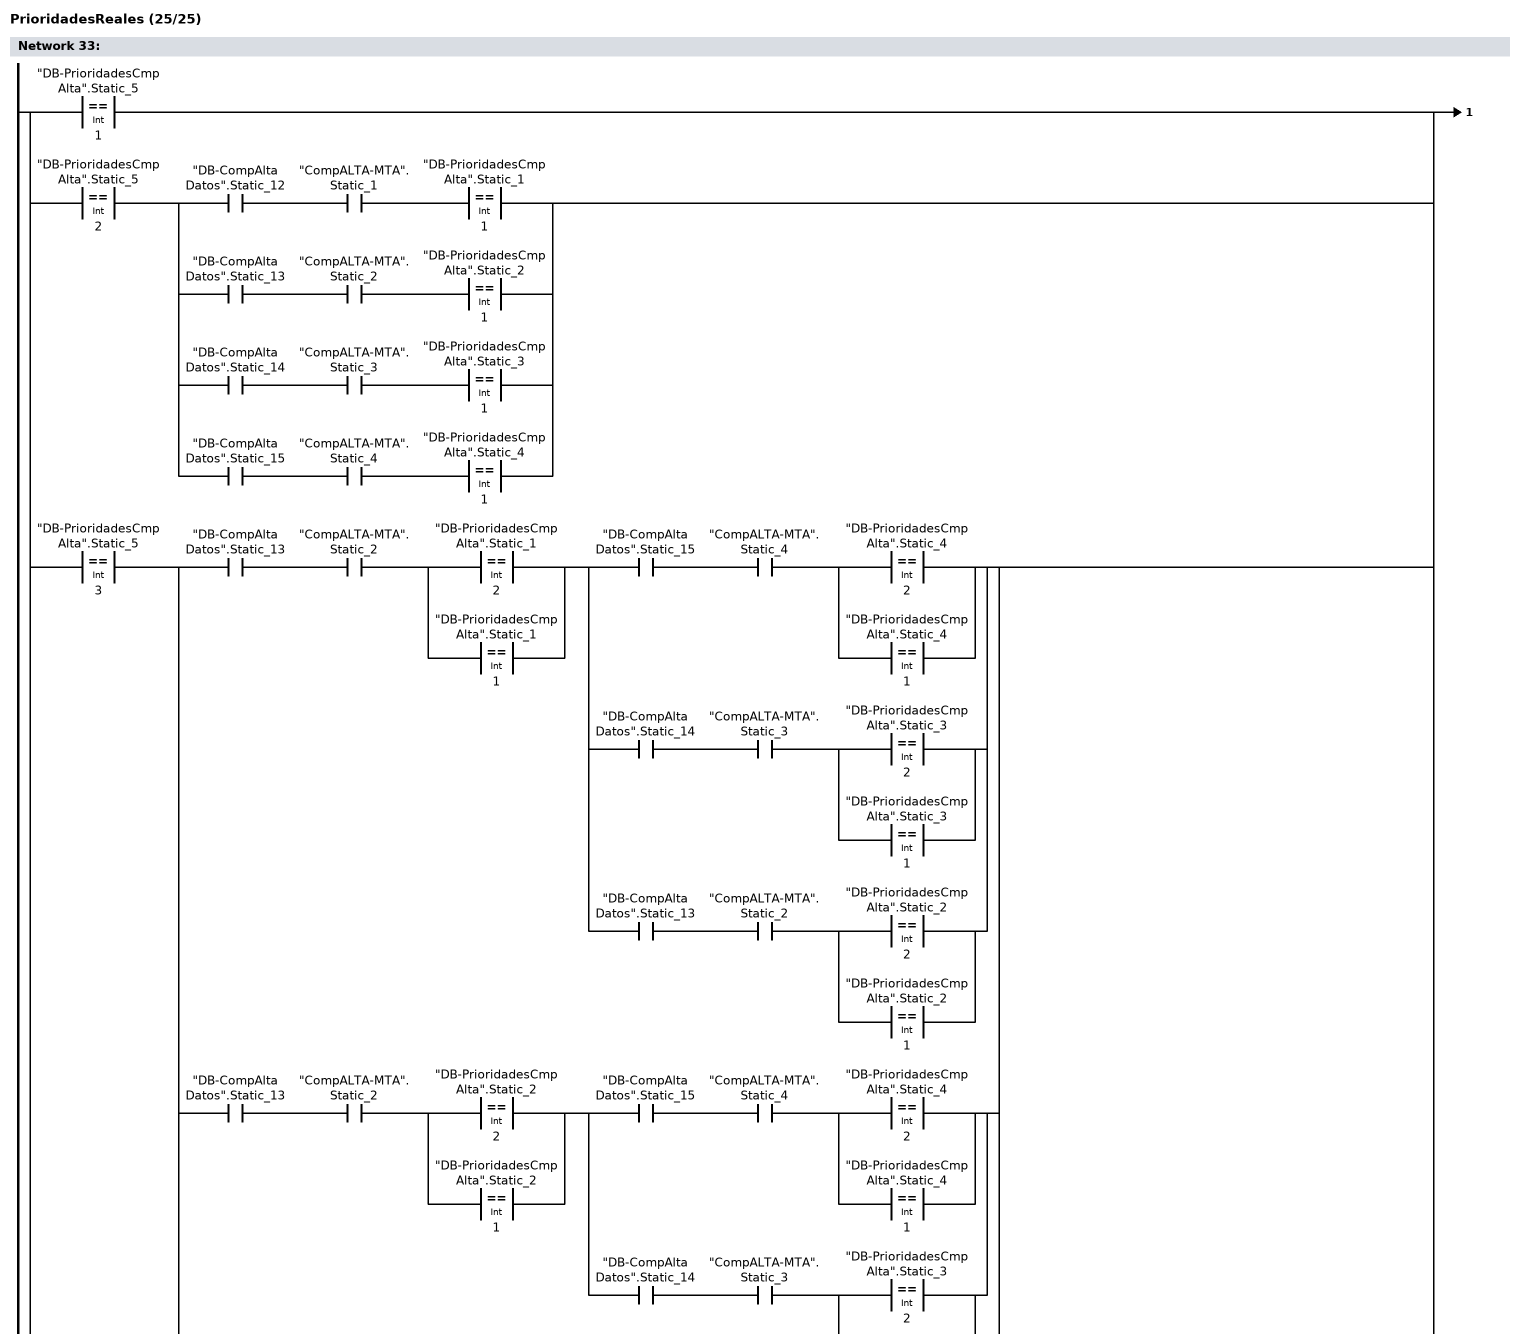
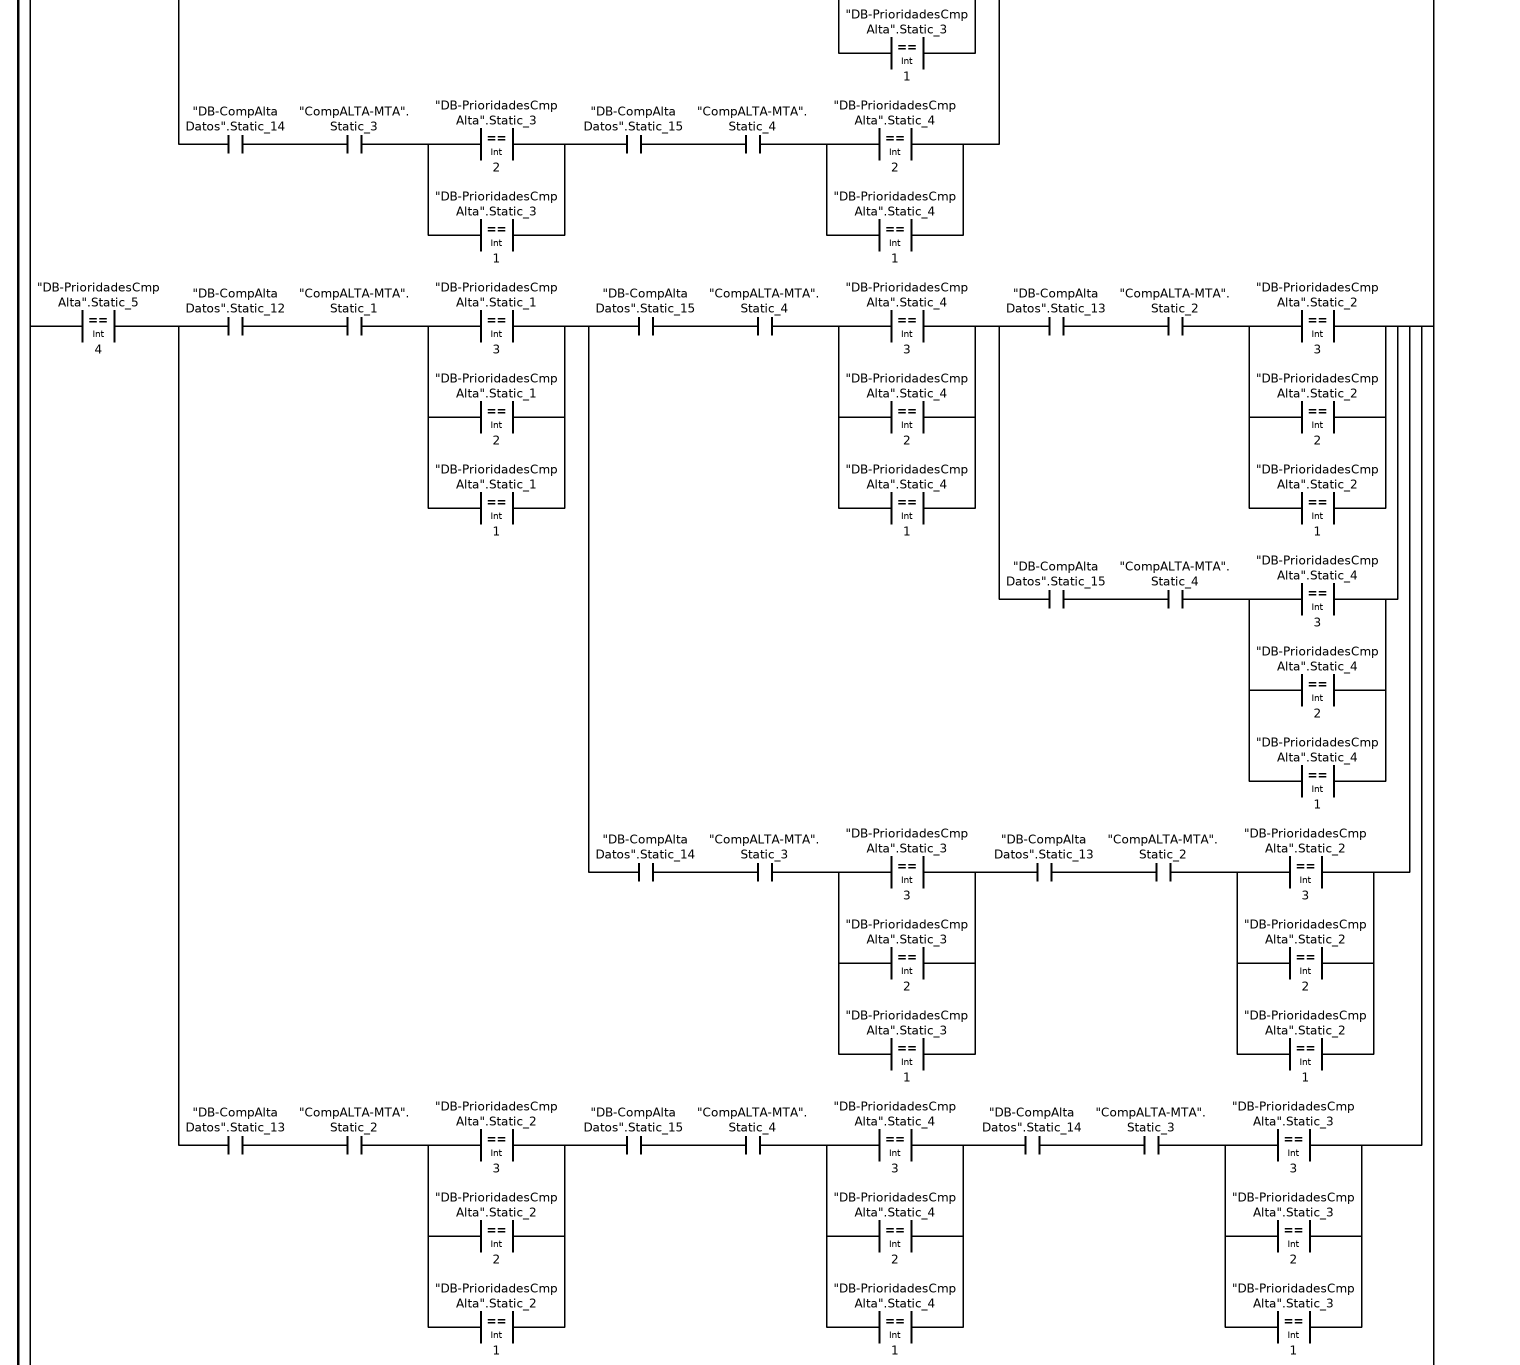
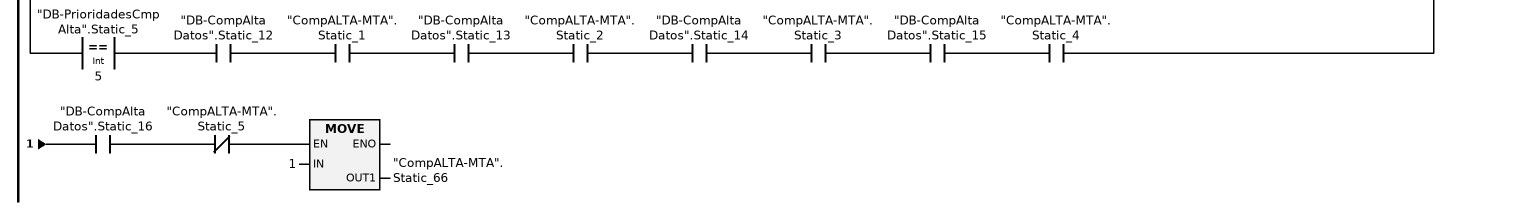
   IF (("DB-PrioridadesCmpAlta".Static_5 = 1) OR (("DB-PrioridadesCmpAlta".Static_5 = 2) AND (("DB-CompAltaDatos".Static_12 AND "CompALTA-MTA".Static_1 AND ("DB-PrioridadesCmpAlta".Static_1 = 1)) OR ("DB-CompAltaDatos".Static_13 AND "CompALTA-MTA".Static_2 AND ("DB-PrioridadesCmpAlta".Static_2 = 1)) OR ("DB-CompAltaDatos".Static_14 AND "CompALTA-MTA".Static_3 AND ("DB-PrioridadesCmpAlta".Static_3 = 1)) OR ("DB-CompAltaDatos".Static_15 AND "CompALTA-MTA".Static_4 AND ("DB-PrioridadesCmpAlta".Static_4 = 1)))) OR (("DB-PrioridadesCmpAlta".Static_5 = 3) AND (("DB-CompAltaDatos".Static_13 AND "CompALTA-MTA".Static_2 AND (("DB-PrioridadesCmpAlta".Static_1 = 2) OR ("DB-PrioridadesCmpAlta".Static_1 = 1)) AND (("DB-CompAltaDatos".Static_15 AND "CompALTA-MTA".Static_4 AND (("DB-PrioridadesCmpAlta".Static_4 = 2) OR ("DB-PrioridadesCmpAlta".Static_4 = 1))) OR ("DB-CompAltaDatos".Static_14 AND "CompALTA-MTA".Static_3 AND (("DB-PrioridadesCmpAlta".Static_3 = 2) OR ("DB-PrioridadesCmpAlta".Static_3 = 1))) OR ("DB-CompAltaDatos".Static_13 AND "CompALTA-MTA".Static_2 AND (("DB-PrioridadesCmpAlta".Static_2 = 2) OR ("DB-PrioridadesCmpAlta".Static_2 = 1))))) OR ("DB-CompAltaDatos".Static_13 AND "CompALTA-MTA".Static_2 AND (("DB-PrioridadesCmpAlta".Static_2 = 2) OR ("DB-PrioridadesCmpAlta".Static_2 = 1)) AND (("DB-CompAltaDatos".Static_15 AND "CompALTA-MTA".Static_4 AND (("DB-PrioridadesCmpAlta".Static_4 = 2) OR ("DB-PrioridadesCmpAlta".Static_4 = 1))) OR ("DB-CompAltaDatos".Static_14 AND "CompALTA-MTA".Static_3 AND (("DB-PrioridadesCmpAlta".Static_3 = 2) OR ("DB-PrioridadesCmpAlta".Static_3 = 1))))) OR ("DB-CompAltaDatos".Static_14 AND "CompALTA-MTA".Static_3 AND (("DB-PrioridadesCmpAlta".Static_3 = 2) OR ("DB-PrioridadesCmpAlta".Static_3 = 1)) AND "DB-CompAltaDatos".Static_15 AND "CompALTA-MTA".Static_4 AND (("DB-PrioridadesCmpAlta".Static_4 = 2) OR ("DB-PrioridadesCmpAlta".Static_4 = 1))))) OR (("DB-PrioridadesCmpAlta".Static_5 = 4) AND (("DB-CompAltaDatos".Static_12 AND "CompALTA-MTA".Static_1 AND (("DB-PrioridadesCmpAlta".Static_1 = 3) OR ("DB-PrioridadesCmpAlta".Static_1 = 2) OR ("DB-PrioridadesCmpAlta".Static_1 = 1)) AND (("DB-CompAltaDatos".Static_15 AND "CompALTA-MTA".Static_4 AND (("DB-PrioridadesCmpAlta".Static_4 = 3) OR ("DB-PrioridadesCmpAlta".Static_4 = 2) OR ("DB-PrioridadesCmpAlta".Static_4 = 1)) AND (("DB-CompAltaDatos".Static_13 AND "CompALTA-MTA".Static_2 AND (("DB-PrioridadesCmpAlta".Static_2 = 3) OR ("DB-PrioridadesCmpAlta".Static_2 = 2) OR ("DB-PrioridadesCmpAlta".Static_2 = 1))) OR ("DB-CompAltaDatos".Static_15 AND "CompALTA-MTA".Static_4 AND (("DB-PrioridadesCmpAlta".Static_4 = 3) OR ("DB-PrioridadesCmpAlta".Static_4 = 2) OR ("DB-PrioridadesCmpAlta".Static_4 = 1))))) OR ("DB-CompAltaDatos".Static_14 AND "CompALTA-MTA".Static_3 AND (("DB-PrioridadesCmpAlta".Static_3 = 3) OR ("DB-PrioridadesCmpAlta".Static_3 = 2) OR ("DB-PrioridadesCmpAlta".Static_3 = 1)) AND "DB-CompAltaDatos".Static_13 AND "CompALTA-MTA".Static_2 AND (("DB-PrioridadesCmpAlta".Static_2 = 3) OR ("DB-PrioridadesCmpAlta".Static_2 = 2) OR ("DB-PrioridadesCmpAlta".Static_2 = 1))))) OR ("DB-CompAltaDatos".Static_13 AND "CompALTA-MTA".Static_2 AND (("DB-PrioridadesCmpAlta".Static_2 = 3) OR ("DB-PrioridadesCmpAlta".Static_2 = 2) OR ("DB-PrioridadesCmpAlta".Static_2 = 1)) AND "DB-CompAltaDatos".Static_15 AND "CompALTA-MTA".Static_4 AND (("DB-PrioridadesCmpAlta".Static_4 = 3) OR ("DB-PrioridadesCmpAlta".Static_4 = 2) OR ("DB-PrioridadesCmpAlta".Static_4 = 1)) AND "DB-CompAltaDatos".Static_14 AND "CompALTA-MTA".Static_3 AND (("DB-PrioridadesCmpAlta".Static_3 = 3) OR ("DB-PrioridadesCmpAlta".Static_3 = 2) OR ("DB-PrioridadesCmpAlta".Static_3 = 1))))) OR (("DB-PrioridadesCmpAlta".Static_5 = 5) AND "DB-CompAltaDatos".Static_12 AND "CompALTA-MTA".Static_1 AND "DB-CompAltaDatos".Static_13 AND "CompALTA-MTA".Static_2 AND "DB-CompAltaDatos".Static_14 AND "CompALTA-MTA".Static_3 AND "DB-CompAltaDatos".Static_15 AND "CompALTA-MTA".Static_4)) AND "DB-CompAltaDatos".Static_16 AND NOT "CompALTA-MTA".Static_5 THEN
       "CompALTA-MTA".Static_66 := 1;
   END_IF;
END_REGION
END_FUNCTION

FUNCTION "FlancosCmpAlta" : Void   // FC45, LAD
{ S7_Optimized_Access := 'FALSE' }
VERSION : 0.1
   VAR_TEMP   // added for the SCL form of the ladder/FBD networks
      _w1 : Bool;
      _w2 : Bool;
      _w3 : Bool;
      _w4 : Bool;
      _w5 : Bool;
      _w6 : Bool;
      _w7 : Bool;
      _s5time1 : S5Time;
   END_VAR
BEGIN

REGION Network 1
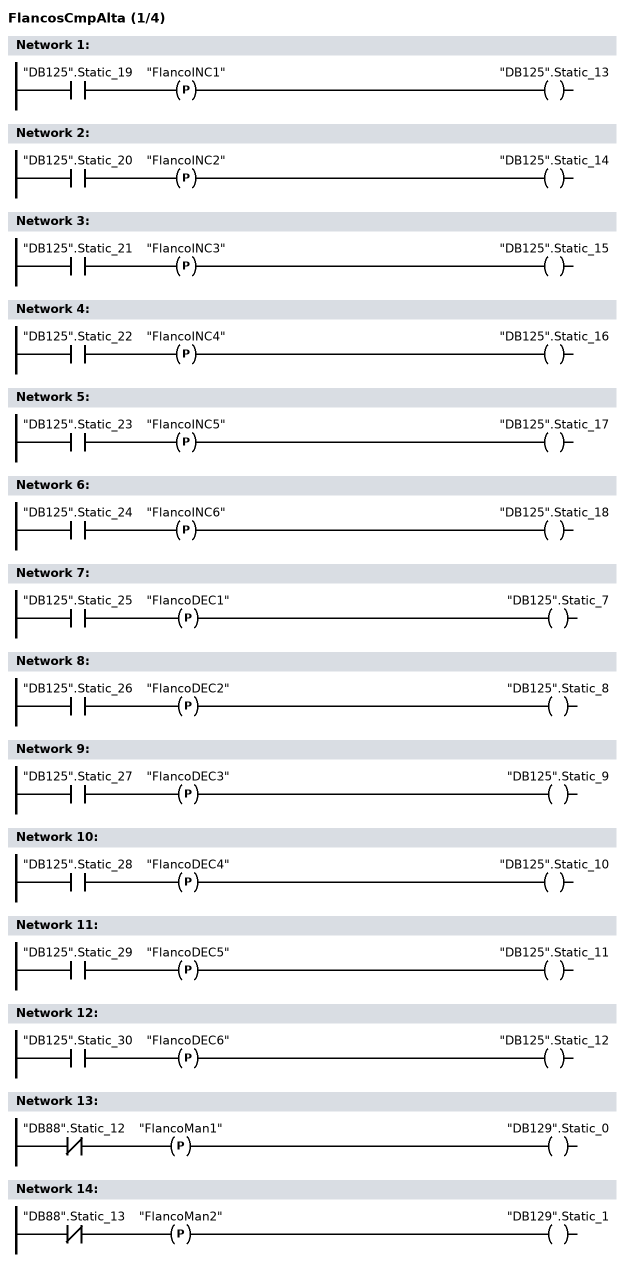
   RUNG wire#powerrail
      Contact( "DB125".Static_19 )
      P_Trig( "FlancoINC1" )
      Coil( "DB125".Static_13 )
   END_RUNG
   // the same network as SCL:
   #_w1 := "DB125".Static_19 AND NOT "FlancoINC1";   // rising edge
   "FlancoINC1" := "DB125".Static_19;
   "DB125".Static_13 := #_w1;
END_REGION

REGION Network 2
   RUNG wire#powerrail
      Contact( "DB125".Static_20 )
      P_Trig( "FlancoINC2" )
      Coil( "DB125".Static_14 )
   END_RUNG
   // the same network as SCL:
   #_w1 := "DB125".Static_20 AND NOT "FlancoINC2";   // rising edge
   "FlancoINC2" := "DB125".Static_20;
   "DB125".Static_14 := #_w1;
END_REGION

REGION Network 3
   RUNG wire#powerrail
      Contact( "DB125".Static_21 )
      P_Trig( "FlancoINC3" )
      Coil( "DB125".Static_15 )
   END_RUNG
   // the same network as SCL:
   #_w1 := "DB125".Static_21 AND NOT "FlancoINC3";   // rising edge
   "FlancoINC3" := "DB125".Static_21;
   "DB125".Static_15 := #_w1;
END_REGION

REGION Network 4
   RUNG wire#powerrail
      Contact( "DB125".Static_22 )
      P_Trig( "FlancoINC4" )
      Coil( "DB125".Static_16 )
   END_RUNG
   // the same network as SCL:
   #_w1 := "DB125".Static_22 AND NOT "FlancoINC4";   // rising edge
   "FlancoINC4" := "DB125".Static_22;
   "DB125".Static_16 := #_w1;
END_REGION

REGION Network 5
   RUNG wire#powerrail
      Contact( "DB125".Static_23 )
      P_Trig( "FlancoINC5" )
      Coil( "DB125".Static_17 )
   END_RUNG
   // the same network as SCL:
   #_w1 := "DB125".Static_23 AND NOT "FlancoINC5";   // rising edge
   "FlancoINC5" := "DB125".Static_23;
   "DB125".Static_17 := #_w1;
END_REGION

REGION Network 6
   RUNG wire#powerrail
      Contact( "DB125".Static_24 )
      P_Trig( "FlancoINC6" )
      Coil( "DB125".Static_18 )
   END_RUNG
   // the same network as SCL:
   #_w1 := "DB125".Static_24 AND NOT "FlancoINC6";   // rising edge
   "FlancoINC6" := "DB125".Static_24;
   "DB125".Static_18 := #_w1;
END_REGION

REGION Network 7
   RUNG wire#powerrail
      Contact( "DB125".Static_25 )
      P_Trig( "FlancoDEC1" )
      Coil( "DB125".Static_7 )
   END_RUNG
   // the same network as SCL:
   #_w1 := "DB125".Static_25 AND NOT "FlancoDEC1";   // rising edge
   "FlancoDEC1" := "DB125".Static_25;
   "DB125".Static_7 := #_w1;
END_REGION

REGION Network 8
   RUNG wire#powerrail
      Contact( "DB125".Static_26 )
      P_Trig( "FlancoDEC2" )
      Coil( "DB125".Static_8 )
   END_RUNG
   // the same network as SCL:
   #_w1 := "DB125".Static_26 AND NOT "FlancoDEC2";   // rising edge
   "FlancoDEC2" := "DB125".Static_26;
   "DB125".Static_8 := #_w1;
END_REGION

REGION Network 9
   RUNG wire#powerrail
      Contact( "DB125".Static_27 )
      P_Trig( "FlancoDEC3" )
      Coil( "DB125".Static_9 )
   END_RUNG
   // the same network as SCL:
   #_w1 := "DB125".Static_27 AND NOT "FlancoDEC3";   // rising edge
   "FlancoDEC3" := "DB125".Static_27;
   "DB125".Static_9 := #_w1;
END_REGION

REGION Network 10
   RUNG wire#powerrail
      Contact( "DB125".Static_28 )
      P_Trig( "FlancoDEC4" )
      Coil( "DB125".Static_10 )
   END_RUNG
   // the same network as SCL:
   #_w1 := "DB125".Static_28 AND NOT "FlancoDEC4";   // rising edge
   "FlancoDEC4" := "DB125".Static_28;
   "DB125".Static_10 := #_w1;
END_REGION

REGION Network 11
   RUNG wire#powerrail
      Contact( "DB125".Static_29 )
      P_Trig( "FlancoDEC5" )
      Coil( "DB125".Static_11 )
   END_RUNG
   // the same network as SCL:
   #_w1 := "DB125".Static_29 AND NOT "FlancoDEC5";   // rising edge
   "FlancoDEC5" := "DB125".Static_29;
   "DB125".Static_11 := #_w1;
END_REGION

REGION Network 12
   RUNG wire#powerrail
      Contact( "DB125".Static_30 )
      P_Trig( "FlancoDEC6" )
      Coil( "DB125".Static_12 )
   END_RUNG
   // the same network as SCL:
   #_w1 := "DB125".Static_30 AND NOT "FlancoDEC6";   // rising edge
   "FlancoDEC6" := "DB125".Static_30;
   "DB125".Static_12 := #_w1;
END_REGION

REGION Network 13
   RUNG wire#powerrail
      I_Contact( "DB88".Static_12 )
      P_Trig( "FlancoMan1" )
      Coil( "DB129".Static_0 )
   END_RUNG
   // the same network as SCL:
   #_w1 := NOT "DB88".Static_12 AND NOT "FlancoMan1";   // rising edge
   "FlancoMan1" := NOT "DB88".Static_12;
   "DB129".Static_0 := #_w1;
END_REGION

REGION Network 14
   RUNG wire#powerrail
      I_Contact( "DB88".Static_13 )
      P_Trig( "FlancoMan2" )
      Coil( "DB129".Static_1 )
   END_RUNG
   // the same network as SCL:
   #_w1 := NOT "DB88".Static_13 AND NOT "FlancoMan2";   // rising edge
   "FlancoMan2" := NOT "DB88".Static_13;
   "DB129".Static_1 := #_w1;
END_REGION

REGION Network 15
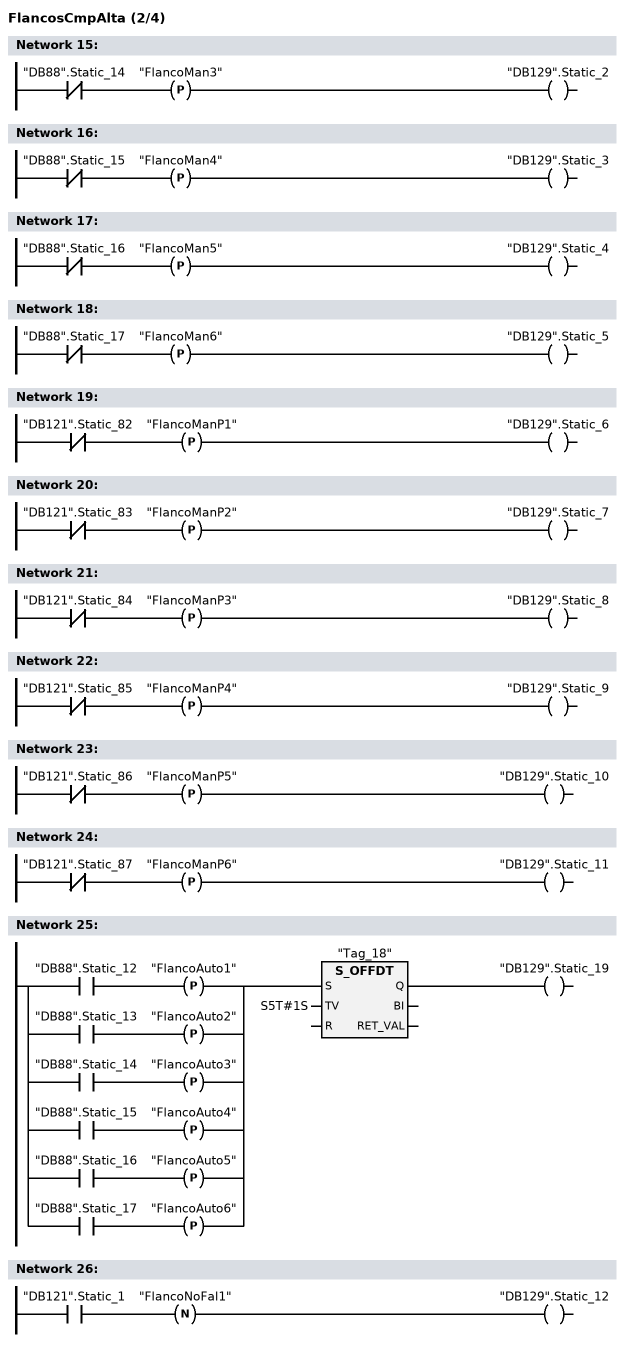
   RUNG wire#powerrail
      I_Contact( "DB88".Static_14 )
      P_Trig( "FlancoMan3" )
      Coil( "DB129".Static_2 )
   END_RUNG
   // the same network as SCL:
   #_w1 := NOT "DB88".Static_14 AND NOT "FlancoMan3";   // rising edge
   "FlancoMan3" := NOT "DB88".Static_14;
   "DB129".Static_2 := #_w1;
END_REGION

REGION Network 16
   RUNG wire#powerrail
      I_Contact( "DB88".Static_15 )
      P_Trig( "FlancoMan4" )
      Coil( "DB129".Static_3 )
   END_RUNG
   // the same network as SCL:
   #_w1 := NOT "DB88".Static_15 AND NOT "FlancoMan4";   // rising edge
   "FlancoMan4" := NOT "DB88".Static_15;
   "DB129".Static_3 := #_w1;
END_REGION

REGION Network 17
   RUNG wire#powerrail
      I_Contact( "DB88".Static_16 )
      P_Trig( "FlancoMan5" )
      Coil( "DB129".Static_4 )
   END_RUNG
   // the same network as SCL:
   #_w1 := NOT "DB88".Static_16 AND NOT "FlancoMan5";   // rising edge
   "FlancoMan5" := NOT "DB88".Static_16;
   "DB129".Static_4 := #_w1;
END_REGION

REGION Network 18
   RUNG wire#powerrail
      I_Contact( "DB88".Static_17 )
      P_Trig( "FlancoMan6" )
      Coil( "DB129".Static_5 )
   END_RUNG
   // the same network as SCL:
   #_w1 := NOT "DB88".Static_17 AND NOT "FlancoMan6";   // rising edge
   "FlancoMan6" := NOT "DB88".Static_17;
   "DB129".Static_5 := #_w1;
END_REGION

REGION Network 19
   RUNG wire#powerrail
      I_Contact( "DB121".Static_82 )
      P_Trig( "FlancoManP1" )
      Coil( "DB129".Static_6 )
   END_RUNG
   // the same network as SCL:
   #_w1 := NOT "DB121".Static_82 AND NOT "FlancoManP1";   // rising edge
   "FlancoManP1" := NOT "DB121".Static_82;
   "DB129".Static_6 := #_w1;
END_REGION

REGION Network 20
   RUNG wire#powerrail
      I_Contact( "DB121".Static_83 )
      P_Trig( "FlancoManP2" )
      Coil( "DB129".Static_7 )
   END_RUNG
   // the same network as SCL:
   #_w1 := NOT "DB121".Static_83 AND NOT "FlancoManP2";   // rising edge
   "FlancoManP2" := NOT "DB121".Static_83;
   "DB129".Static_7 := #_w1;
END_REGION

REGION Network 21
   RUNG wire#powerrail
      I_Contact( "DB121".Static_84 )
      P_Trig( "FlancoManP3" )
      Coil( "DB129".Static_8 )
   END_RUNG
   // the same network as SCL:
   #_w1 := NOT "DB121".Static_84 AND NOT "FlancoManP3";   // rising edge
   "FlancoManP3" := NOT "DB121".Static_84;
   "DB129".Static_8 := #_w1;
END_REGION

REGION Network 22
   RUNG wire#powerrail
      I_Contact( "DB121".Static_85 )
      P_Trig( "FlancoManP4" )
      Coil( "DB129".Static_9 )
   END_RUNG
   // the same network as SCL:
   #_w1 := NOT "DB121".Static_85 AND NOT "FlancoManP4";   // rising edge
   "FlancoManP4" := NOT "DB121".Static_85;
   "DB129".Static_9 := #_w1;
END_REGION

REGION Network 23
   RUNG wire#powerrail
      I_Contact( "DB121".Static_86 )
      P_Trig( "FlancoManP5" )
      Coil( "DB129".Static_10 )
   END_RUNG
   // the same network as SCL:
   #_w1 := NOT "DB121".Static_86 AND NOT "FlancoManP5";   // rising edge
   "FlancoManP5" := NOT "DB121".Static_86;
   "DB129".Static_10 := #_w1;
END_REGION

REGION Network 24
   RUNG wire#powerrail
      I_Contact( "DB121".Static_87 )
      P_Trig( "FlancoManP6" )
      Coil( "DB129".Static_11 )
   END_RUNG
   // the same network as SCL:
   #_w1 := NOT "DB121".Static_87 AND NOT "FlancoManP6";   // rising edge
   "FlancoManP6" := NOT "DB121".Static_87;
   "DB129".Static_11 := #_w1;
END_REGION

REGION Network 25
   RUNG wire#powerrail
      Contact( "DB88".Static_12 )
      P_Trig( "FlancoAuto1" )
      wire#w1
      S_OFFDT(T_NO := "Tag_18", TV := S5T#1S, R :=, BI =>, RET_VAL =>)
      Coil( "DB129".Static_19 )
   END_RUNG
   RUNG wire#powerrail
      Contact( "DB88".Static_13 )
      P_Trig( "FlancoAuto2" )
   END_RUNG wire#w1
   RUNG wire#powerrail
      Contact( "DB88".Static_14 )
      P_Trig( "FlancoAuto3" )
   END_RUNG wire#w1
   RUNG wire#powerrail
      Contact( "DB88".Static_15 )
      P_Trig( "FlancoAuto4" )
   END_RUNG wire#w1
   RUNG wire#powerrail
      Contact( "DB88".Static_16 )
      P_Trig( "FlancoAuto5" )
   END_RUNG wire#w1
   RUNG wire#powerrail
      Contact( "DB88".Static_17 )
      P_Trig( "FlancoAuto6" )
   END_RUNG wire#w1
   // the same network as SCL:
   #_w1 := "DB88".Static_12 AND NOT "FlancoAuto1";   // rising edge
   "FlancoAuto1" := "DB88".Static_12;
   #_w2 := "DB88".Static_13 AND NOT "FlancoAuto2";   // rising edge
   "FlancoAuto2" := "DB88".Static_13;
   #_w3 := "DB88".Static_14 AND NOT "FlancoAuto3";   // rising edge
   "FlancoAuto3" := "DB88".Static_14;
   #_w4 := "DB88".Static_15 AND NOT "FlancoAuto4";   // rising edge
   "FlancoAuto4" := "DB88".Static_15;
   #_w5 := "DB88".Static_16 AND NOT "FlancoAuto5";   // rising edge
   "FlancoAuto5" := "DB88".Static_16;
   #_w6 := "DB88".Static_17 AND NOT "FlancoAuto6";   // rising edge
   "FlancoAuto6" := "DB88".Static_17;
   #_s5time1 := S_OFFDT(T_NO := "Tag_18",
                        S := #_w1 OR #_w2 OR #_w3 OR #_w4 OR #_w5 OR #_w6,
                        TV := S5T#1S,
                        Q => #_w7);
   "DB129".Static_19 := #_w7;
END_REGION

REGION Network 26
   RUNG wire#powerrail
      Contact( "DB121".Static_1 )
      N_Trig( "FlancoNoFal1" )
      Coil( "DB129".Static_12 )
   END_RUNG
   // the same network as SCL:
   #_w1 := NOT "DB121".Static_1 AND "FlancoNoFal1";   // falling edge
   "FlancoNoFal1" := "DB121".Static_1;
   "DB129".Static_12 := #_w1;
END_REGION

REGION Network 27
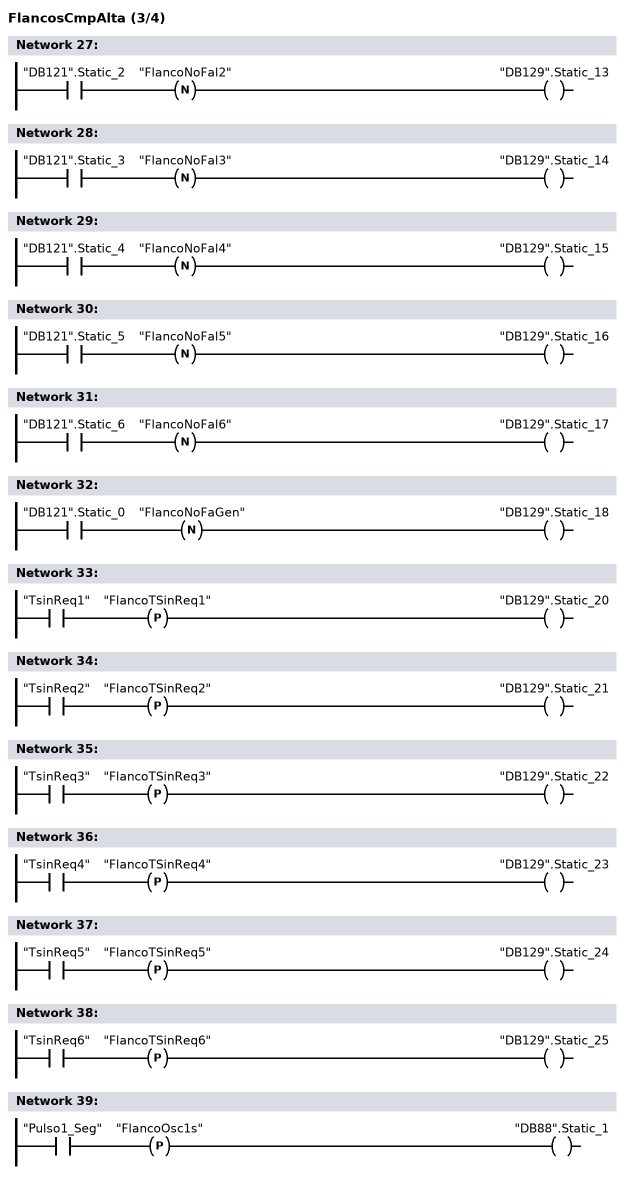
   RUNG wire#powerrail
      Contact( "DB121".Static_2 )
      N_Trig( "FlancoNoFal2" )
      Coil( "DB129".Static_13 )
   END_RUNG
   // the same network as SCL:
   #_w1 := NOT "DB121".Static_2 AND "FlancoNoFal2";   // falling edge
   "FlancoNoFal2" := "DB121".Static_2;
   "DB129".Static_13 := #_w1;
END_REGION

REGION Network 28
   RUNG wire#powerrail
      Contact( "DB121".Static_3 )
      N_Trig( "FlancoNoFal3" )
      Coil( "DB129".Static_14 )
   END_RUNG
   // the same network as SCL:
   #_w1 := NOT "DB121".Static_3 AND "FlancoNoFal3";   // falling edge
   "FlancoNoFal3" := "DB121".Static_3;
   "DB129".Static_14 := #_w1;
END_REGION

REGION Network 29
   RUNG wire#powerrail
      Contact( "DB121".Static_4 )
      N_Trig( "FlancoNoFal4" )
      Coil( "DB129".Static_15 )
   END_RUNG
   // the same network as SCL:
   #_w1 := NOT "DB121".Static_4 AND "FlancoNoFal4";   // falling edge
   "FlancoNoFal4" := "DB121".Static_4;
   "DB129".Static_15 := #_w1;
END_REGION

REGION Network 30
   RUNG wire#powerrail
      Contact( "DB121".Static_5 )
      N_Trig( "FlancoNoFal5" )
      Coil( "DB129".Static_16 )
   END_RUNG
   // the same network as SCL:
   #_w1 := NOT "DB121".Static_5 AND "FlancoNoFal5";   // falling edge
   "FlancoNoFal5" := "DB121".Static_5;
   "DB129".Static_16 := #_w1;
END_REGION

REGION Network 31
   RUNG wire#powerrail
      Contact( "DB121".Static_6 )
      N_Trig( "FlancoNoFal6" )
      Coil( "DB129".Static_17 )
   END_RUNG
   // the same network as SCL:
   #_w1 := NOT "DB121".Static_6 AND "FlancoNoFal6";   // falling edge
   "FlancoNoFal6" := "DB121".Static_6;
   "DB129".Static_17 := #_w1;
END_REGION

REGION Network 32
   RUNG wire#powerrail
      Contact( "DB121".Static_0 )
      N_Trig( "FlancoNoFaGen" )
      Coil( "DB129".Static_18 )
   END_RUNG
   // the same network as SCL:
   #_w1 := NOT "DB121".Static_0 AND "FlancoNoFaGen";   // falling edge
   "FlancoNoFaGen" := "DB121".Static_0;
   "DB129".Static_18 := #_w1;
END_REGION

REGION Network 33
   RUNG wire#powerrail
      Contact( "TsinReq1" )
      P_Trig( "FlancoTSinReq1" )
      Coil( "DB129".Static_20 )
   END_RUNG
   // the same network as SCL:
   #_w1 := "TsinReq1" AND NOT "FlancoTSinReq1";   // rising edge
   "FlancoTSinReq1" := "TsinReq1";
   "DB129".Static_20 := #_w1;
END_REGION

REGION Network 34
   RUNG wire#powerrail
      Contact( "TsinReq2" )
      P_Trig( "FlancoTSinReq2" )
      Coil( "DB129".Static_21 )
   END_RUNG
   // the same network as SCL:
   #_w1 := "TsinReq2" AND NOT "FlancoTSinReq2";   // rising edge
   "FlancoTSinReq2" := "TsinReq2";
   "DB129".Static_21 := #_w1;
END_REGION

REGION Network 35
   RUNG wire#powerrail
      Contact( "TsinReq3" )
      P_Trig( "FlancoTSinReq3" )
      Coil( "DB129".Static_22 )
   END_RUNG
   // the same network as SCL:
   #_w1 := "TsinReq3" AND NOT "FlancoTSinReq3";   // rising edge
   "FlancoTSinReq3" := "TsinReq3";
   "DB129".Static_22 := #_w1;
END_REGION

REGION Network 36
   RUNG wire#powerrail
      Contact( "TsinReq4" )
      P_Trig( "FlancoTSinReq4" )
      Coil( "DB129".Static_23 )
   END_RUNG
   // the same network as SCL:
   #_w1 := "TsinReq4" AND NOT "FlancoTSinReq4";   // rising edge
   "FlancoTSinReq4" := "TsinReq4";
   "DB129".Static_23 := #_w1;
END_REGION

REGION Network 37
   RUNG wire#powerrail
      Contact( "TsinReq5" )
      P_Trig( "FlancoTSinReq5" )
      Coil( "DB129".Static_24 )
   END_RUNG
   // the same network as SCL:
   #_w1 := "TsinReq5" AND NOT "FlancoTSinReq5";   // rising edge
   "FlancoTSinReq5" := "TsinReq5";
   "DB129".Static_24 := #_w1;
END_REGION

REGION Network 38
   RUNG wire#powerrail
      Contact( "TsinReq6" )
      P_Trig( "FlancoTSinReq6" )
      Coil( "DB129".Static_25 )
   END_RUNG
   // the same network as SCL:
   #_w1 := "TsinReq6" AND NOT "FlancoTSinReq6";   // rising edge
   "FlancoTSinReq6" := "TsinReq6";
   "DB129".Static_25 := #_w1;
END_REGION

REGION Network 39
   RUNG wire#powerrail
      Contact( "Pulso1_Seg" )
      P_Trig( "FlancoOsc1s" )
      Coil( "DB88".Static_1 )
   END_RUNG
   // the same network as SCL:
   #_w1 := "Pulso1_Seg" AND NOT "FlancoOsc1s";   // rising edge
   "FlancoOsc1s" := "Pulso1_Seg";
   "DB88".Static_1 := #_w1;
END_REGION

REGION Network 40
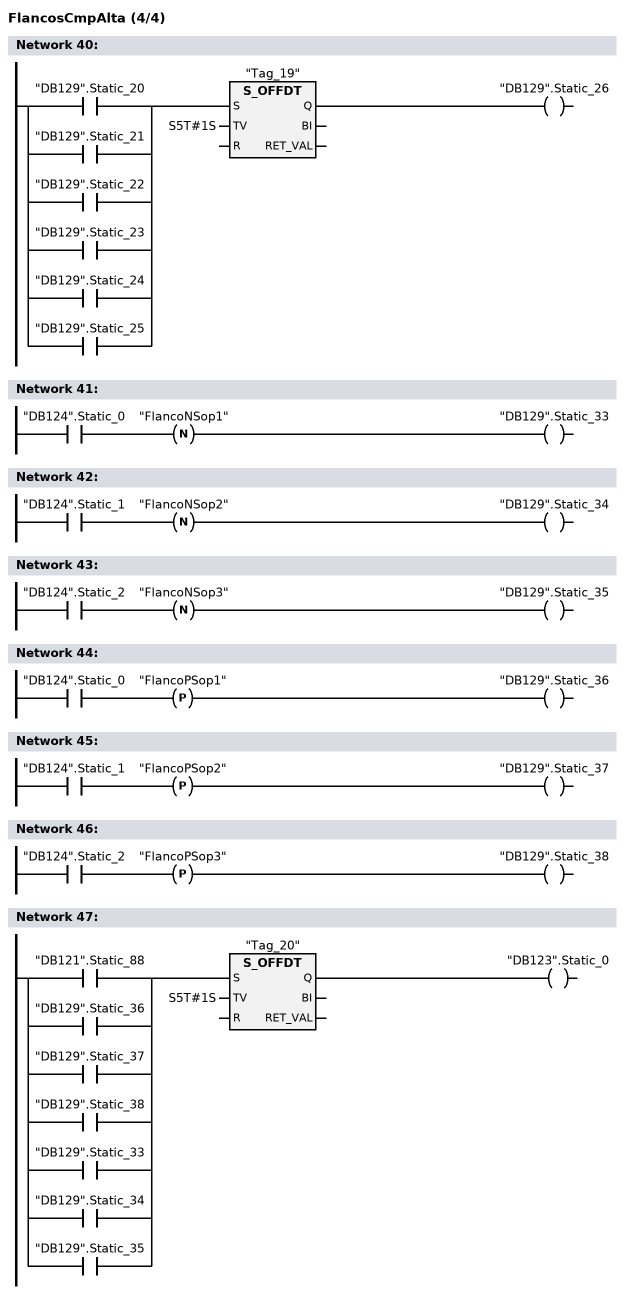
   RUNG wire#powerrail
      Contact( "DB129".Static_20 )
      wire#w1
      S_OFFDT(T_NO := "Tag_19", TV := S5T#1S, R :=, BI =>, RET_VAL =>)
      Coil( "DB129".Static_26 )
   END_RUNG
   RUNG wire#powerrail
      Contact( "DB129".Static_21 )
   END_RUNG wire#w1
   RUNG wire#powerrail
      Contact( "DB129".Static_22 )
   END_RUNG wire#w1
   RUNG wire#powerrail
      Contact( "DB129".Static_23 )
   END_RUNG wire#w1
   RUNG wire#powerrail
      Contact( "DB129".Static_24 )
   END_RUNG wire#w1
   RUNG wire#powerrail
      Contact( "DB129".Static_25 )
   END_RUNG wire#w1
   // the same network as SCL:
   #_s5time1 := S_OFFDT(T_NO := "Tag_19",
                        S := "DB129".Static_20 OR "DB129".Static_21 OR "DB129".Static_22 OR "DB129".Static_23 OR "DB129".Static_24 OR "DB129".Static_25,
                        TV := S5T#1S,
                        Q => #_w1);
   "DB129".Static_26 := #_w1;
END_REGION

REGION Network 41
   RUNG wire#powerrail
      Contact( "DB124".Static_0 )
      N_Trig( "FlancoNSop1" )
      Coil( "DB129".Static_33 )
   END_RUNG
   // the same network as SCL:
   #_w1 := NOT "DB124".Static_0 AND "FlancoNSop1";   // falling edge
   "FlancoNSop1" := "DB124".Static_0;
   "DB129".Static_33 := #_w1;
END_REGION

REGION Network 42
   RUNG wire#powerrail
      Contact( "DB124".Static_1 )
      N_Trig( "FlancoNSop2" )
      Coil( "DB129".Static_34 )
   END_RUNG
   // the same network as SCL:
   #_w1 := NOT "DB124".Static_1 AND "FlancoNSop2";   // falling edge
   "FlancoNSop2" := "DB124".Static_1;
   "DB129".Static_34 := #_w1;
END_REGION

REGION Network 43
   RUNG wire#powerrail
      Contact( "DB124".Static_2 )
      N_Trig( "FlancoNSop3" )
      Coil( "DB129".Static_35 )
   END_RUNG
   // the same network as SCL:
   #_w1 := NOT "DB124".Static_2 AND "FlancoNSop3";   // falling edge
   "FlancoNSop3" := "DB124".Static_2;
   "DB129".Static_35 := #_w1;
END_REGION

REGION Network 44
   RUNG wire#powerrail
      Contact( "DB124".Static_0 )
      P_Trig( "FlancoPSop1" )
      Coil( "DB129".Static_36 )
   END_RUNG
   // the same network as SCL:
   #_w1 := "DB124".Static_0 AND NOT "FlancoPSop1";   // rising edge
   "FlancoPSop1" := "DB124".Static_0;
   "DB129".Static_36 := #_w1;
END_REGION

REGION Network 45
   RUNG wire#powerrail
      Contact( "DB124".Static_1 )
      P_Trig( "FlancoPSop2" )
      Coil( "DB129".Static_37 )
   END_RUNG
   // the same network as SCL:
   #_w1 := "DB124".Static_1 AND NOT "FlancoPSop2";   // rising edge
   "FlancoPSop2" := "DB124".Static_1;
   "DB129".Static_37 := #_w1;
END_REGION

REGION Network 46
   RUNG wire#powerrail
      Contact( "DB124".Static_2 )
      P_Trig( "FlancoPSop3" )
      Coil( "DB129".Static_38 )
   END_RUNG
   // the same network as SCL:
   #_w1 := "DB124".Static_2 AND NOT "FlancoPSop3";   // rising edge
   "FlancoPSop3" := "DB124".Static_2;
   "DB129".Static_38 := #_w1;
END_REGION

REGION Network 47
   RUNG wire#powerrail
      Contact( "DB121".Static_88 )
      wire#w1
      S_OFFDT(T_NO := "Tag_20", TV := S5T#1S, R :=, BI =>, RET_VAL =>)
      Coil( "DB123".Static_0 )
   END_RUNG
   RUNG wire#powerrail
      Contact( "DB129".Static_36 )
   END_RUNG wire#w1
   RUNG wire#powerrail
      Contact( "DB129".Static_37 )
   END_RUNG wire#w1
   RUNG wire#powerrail
      Contact( "DB129".Static_38 )
   END_RUNG wire#w1
   RUNG wire#powerrail
      Contact( "DB129".Static_33 )
   END_RUNG wire#w1
   RUNG wire#powerrail
      Contact( "DB129".Static_34 )
   END_RUNG wire#w1
   RUNG wire#powerrail
      Contact( "DB129".Static_35 )
   END_RUNG wire#w1
   // the same network as SCL:
   #_s5time1 := S_OFFDT(T_NO := "Tag_20",
                        S := "DB121".Static_88 OR "DB129".Static_36 OR "DB129".Static_37 OR "DB129".Static_38 OR "DB129".Static_33 OR "DB129".Static_34 OR "DB129".Static_35,
                        TV := S5T#1S,
                        Q => #_w1);
   "DB123".Static_0 := #_w1;
END_REGION
END_FUNCTION

FUNCTION "CompAltaPanel" : Void   // FC47, LAD
{ S7_Optimized_Access := 'FALSE' }
VERSION : 0.1
   VAR_TEMP   // added for the SCL form of the ladder/FBD networks
      _w1 : Bool;
      _s5time1 : S5Time;
      _w2 : Bool;
   END_VAR
BEGIN

REGION Network 1